// TIA Portal project "TNprojINZ" (V15.1)

(* hardware
DEVICE "S71500/ET200MP station_1"  S7-1500 station
   slot 0: "Rail_0"  Rack  6ES7 590-1***0-0AA0
   slot 1: "PLC_1"  CPU 1516-3 PN/DP  6ES7 516-3AN01-0AB0  V2.5
      slot 3: "CPU display_1"  6ES7591-1BA00-0AA0
   slot 2: "DI 32x24VDC HF_1"  DI 32x24VDC HF  6ES7 521-1BL00-0AB0  V2.1
   slot 3: "DQ 32x24VDC/0.5A ST_1"  DQ 32x24VDC/0.5A ST  6ES7 522-1BL00-0AB0  V2.0
   slot 4: "AI 8xU/I/RTD/TC ST_1"  AI 8xU/I/RTD/TC ST  6ES7 531-7KF00-0AB0  V2.0
   slot 5: "AQ 4xU/I ST_1"  AQ 4xU/I ST  6ES7 532-5HD00-0AB0  V2.0
DEVICE "HMI_1"  TP700 Comfort
   slot 0: "HMI_1"  TP700 Comfort  6AV2 124-0GC01-0AX0  15.1.0.0
   slot 1: "HMI_RT_1"  TP700 Comfort  6AV2 124-0GC01-0AX0  15.1.0.0
   slot 5: "HMI_1.IE_CP_1"  PROFINET Interface  15.0.1.0
      slot 1: "PROFINET Interface_1"  PROFINET Interface
         slot 1: "Port_1"  Port
         slot 2: "Port_2"  Port
   slot 7: "HMI_1.MPI/DP_CP_1"  MPI/DP Interface  15.0.1.0
*)

// ===== PLC "PLC_1"  CPU 1516-3 PN/DP =====

VAR_GLOBAL   // PLC tag table "Default tag table"
   "System_Byte" AT %MB1 : Byte;
   "FirstScan" AT %M1.0 : Bool;
   "DiagStatusUpdate" AT %M1.1 : Bool;
   "AlwaysTRUE" AT %M1.2 : Bool;
   "AlwaysFALSE" AT %M1.3 : Bool;
   "Clock_Byte" AT %MB0 : Byte;
   "Clock_10Hz" AT %M0.0 : Bool;
   "Clock_5Hz" AT %M0.1 : Bool;
   "Clock_2.5Hz" AT %M0.2 : Bool;
   "Clock_2Hz" AT %M0.3 : Bool;
   "Clock_1.25Hz" AT %M0.4 : Bool;
   "Clock_1Hz" AT %M0.5 : Bool;
   "Clock_0.625Hz" AT %M0.6 : Bool;
   "Clock_0.5Hz" AT %M0.7 : Bool;
   "Tag_1" AT %C3 : Counter;
END_VAR

DATA_BLOCK "Ster pompami"   // DB1
{ S7_Optimized_Access := 'TRUE' }
VERSION : 0.1
   VAR
      "przegrzana P1" : Bool;
      "przegrzana P2" : Bool;
      "przegrzana P3" : Bool;
      "przegrzana P4" : Bool;
      "przegrzana P5" : Bool;
      "przegrzana P6" : Bool;
      "przegrzana P7" : Bool;
      "przegrzana P8" : Bool;
   END_VAR
BEGIN
END_DATA_BLOCK

DATA_BLOCK "HMI komunikacja"   // DB2
{ S7_Optimized_Access := 'TRUE' }
VERSION : 0.1
   VAR
      "HMI Temp max Z1" : Real;   // zadany w HMI, następna part produktu
      "HMI Temp max Z2" : Real;   // zadany w HMI, następna part produktu
      "HMI Temp max Z3" : Real;   // zadany w HMI, następna part produktu
      "HMI Temp max Z4" : Real;   // zadany w HMI, następna part produktu
      "HMI poziom cieczy Z1" : Real;   // zadany w HMI, następna part produktu
      "HMI poziom cieczy Z2" : Real;   // zadany w HMI, następna part produktu
      "HMI poziom cieczy Z3" : Real;   // zadany w HMI, następna part produktu
      "HMI poziom cieczy Z4" : Real;   // zadany w HMI, następna part produktu
      "Czas utrz T w Z1 (timer)" : Real := 0.0;
      "Czas utrz T w Z2 (timer)" : Real := 0.0;
      "Czas utrz T w Z3 (timer)" : Real := 0.0;
      "Czas utrz T w Z4 (timer)" : Real := 0.0;
      "HMI czas utrz T  Z1" : Real := 0.0;   // zadany w HMI, następna part produktu
      "HMI czas utrz T  Z2" : Real := 0.0;   // zadany w HMI, następna part produktu
      "HMI czas utrz T  Z3" : Real := 0.0;   // zadany w HMI, następna part produktu
      "HMI czas utrz T  Z4" : Real := 0.0;   // zadany w HMI, następna part produktu
      "rura blue P5 i P6" : Bool := 0;
      "rura blue P1 i P2" : Bool := 0;
      "Start/Stop" : Bool := 0;
      "Blokada zmiany par. PRO" : Bool := 0;
   END_VAR
BEGIN
END_DATA_BLOCK

DATA_BLOCK "OPC - z LabVIEW"   // DB3
{ S7_Optimized_Access := 'FALSE' }
VERSION : 0.1
   VAR
      "Temp P1" : Real;
      "Temp P2" : Real;
      "Temp P3" : Real;
      "Temp P4" : Real;
      "Temp P5" : Real;
      "Temp P6" : Real;
      "Temp P7" : Real;
      "Temp P8" : Real;
      "Temp cieczy w zb1" : Real;
      "Temp cieczy w zb2" : Real;
      "Temp cieczy w zb3" : Real;
      "Temp cieczy w zb4" : Real;
      "Poziom zbiornik 1" : Real;
      "Poziom zbiornik 2" : Real;
      "Poziom zbiornik 3" : Real;
      "Poziom zbiornik 4" : Real;
      komTESTz : Bool := 0;
   END_VAR
BEGIN
END_DATA_BLOCK

DATA_BLOCK "OPC - do LabVIEW"   // DB4
{ S7_Optimized_Access := 'FALSE' }
VERSION : 0.1
   VAR
      "PRO Temp max Z1" : Real;   // dla SFC, aktualna partia produktu
      "PRO Temp max Z2" : Real;   // dla SFC, aktualna partia produktu
      "PRO Temp max Z3" : Real;   // dla SFC, aktualna partia produktu
      "PRO Temp max Z4" : Real;   // dla SFC, aktualna partia produktu
      "PRO poziom cieczy Z1" : Real;   // dla SFC, aktualna partia produktu
      "PRO poziom cieczy Z2" : Real;   // dla SFC, aktualna partia produktu
      "PRO poziom cieczy Z3" : Real;   // dla SFC, aktualna partia produktu
      "PRO poziom cieczy Z4" : Real;   // dla SFC, aktualna partia produktu
      "PRO czas utrz T  Z1" : Real := 0.0;   // dla SFC, aktualna partia produktu
      "PRO czas utrz T  Z2" : Real := 0.0;   // dla SFC, aktualna partia produktu
      "PRO czas utrz T  Z3" : Real := 0.0;   // dla SFC, aktualna partia produktu
      "PRO czas utrz T  Z4" : Real := 0.0;   // dla SFC, aktualna partia produktu
      Awaria : Bool := 0;
      "Pompa 1" : Bool := 0;
      "Pompa 2" : Bool := 0;
      "Pompa 3" : Bool := 0;
      "Pompa 4" : Bool := 0;
      "Pompa 5" : Bool := 0;
      "Pompa 6" : Bool := 0;
      "Pompa 7" : Bool := 0;
      "Pompa 8" : Bool := 0;
      "Zawór wlotowy 1" : Bool := 0;
      "Zawór wlotowy 2" : Bool := 0;
      "Zawór wlotowy 3" : Bool := 0;
      "Grzałka 1" : Bool := 0;
      "Grzałka 2" : Bool := 0;
      "Grzałka 3" : Bool := 0;
      "Grzałka 4" : Bool := 0;
      "HMI konserwacja P1" : Bool := 0;
      "HMI konserwacja P2" : Bool := 0;
      "HMI konserwacja P3" : Bool := 0;
      "HMI konserwacja P4" : Bool := 0;
      "HMI konserwacja P5" : Bool := 0;
      "HMI konserwacja P6" : Bool := 0;
      "HMI konserwacja P7" : Bool := 0;
      "HMI konserwacja P8" : Bool := 0;
      "Zawór spustowy Z1" : Bool := 0;
      "Zawór spustowy Z2" : Bool := 0;
      "Zawór spustowy Z3" : Bool := 0;
      "Zawór spustowy Z4" : Bool := 0;
      komTESTdo : Bool := 0;
   END_VAR
BEGIN
END_DATA_BLOCK

DATA_BLOCK "Ster grzałki/zbior"   // DB5
{ S7_Optimized_Access := 'TRUE' }
VERSION : 0.1
   VAR
      HISTgrzałka1 : Bool;
      HISTgrzałka2 : Bool;
      HISTgrzałka3 : Bool;
      HISTgrzałka4 : Bool;
      "Wszystkie zbiorniki puste" : Bool;
      "Z1 opróżniony" : Bool;
      "Z2 opróżniony" : Bool;
      "Z3 opróżniony" : Bool;
   END_VAR
BEGIN
END_DATA_BLOCK

// folder: DB - Instance

DATA_BLOCK "Zbiornik 1_DB"   // DB6
{ S7_Optimized_Access := 'TRUE' }
VERSION : 0.1
// stored: InstanceOfName Zbiornik 1
"Zbiornik 1"
BEGIN
END_DATA_BLOCK

DATA_BLOCK "Zbiornik 2_DB"   // DB15
{ S7_Optimized_Access := 'TRUE' }
VERSION : 0.1
// stored: InstanceOfName Zbiornik 2
"Zbiornik 2"
BEGIN
END_DATA_BLOCK

DATA_BLOCK "Zbiornik 3_DB"   // DB16
{ S7_Optimized_Access := 'TRUE' }
VERSION : 0.1
// stored: InstanceOfName Zbiornik 3
"Zbiornik 3"
BEGIN
END_DATA_BLOCK

DATA_BLOCK "Zbiornik 4_DB"   // DB17
{ S7_Optimized_Access := 'TRUE' }
VERSION : 0.1
// stored: InstanceOfName Zbiornik 4
"Zbiornik 4"
BEGIN
END_DATA_BLOCK

DATA_BLOCK "SCL - Sterowanie pompami_DB"   // DB18
{ S7_Optimized_Access := 'TRUE' }
VERSION : 0.1
// stored: InstanceOfName SCL - Sterowanie pompami
"SCL - Sterowanie pompami"
BEGIN
END_DATA_BLOCK

DATA_BLOCK "SCL - Napełnianie i kontrola_DB"   // DB19
{ S7_Optimized_Access := 'TRUE' }
VERSION : 0.1
// stored: InstanceOfName SCL - Napełnianie i kontrola
"SCL - Napełnianie i kontrola"
BEGIN
END_DATA_BLOCK

DATA_BLOCK "SCL - Grzanie_DB"   // DB20
{ S7_Optimized_Access := 'TRUE' }
VERSION : 0.1
// stored: InstanceOfName SCL - Grzanie
"SCL - Grzanie"
BEGIN
END_DATA_BLOCK

DATA_BLOCK "SCL - Awaria_DB"   // DB21
{ S7_Optimized_Access := 'TRUE' }
VERSION : 0.1
// stored: InstanceOfName SCL - Awaria i zabezpieczenia par.
"SCL - Awaria i zabezpieczenia par."
BEGIN
END_DATA_BLOCK

DATA_BLOCK "FB - pompy_DB"   // DB22
{ S7_Optimized_Access := 'TRUE' }
VERSION : 0.1
// stored: InstanceOfName FB - pompy
"FB - pompy"
BEGIN
END_DATA_BLOCK

DATA_BLOCK "FB - grzałki_DB"   // DB23
{ S7_Optimized_Access := 'TRUE' }
VERSION : 0.1
// stored: InstanceOfName FB - grzałki
"FB - grzałki"
BEGIN
END_DATA_BLOCK

// folder: System blocks/Program resources

DATA_BLOCK "IEC_Timer_2_DB"   // DB7
{ S7_Optimized_Access := 'TRUE' }
AUTHOR : Simatic
FAMILY : IEC
NAME : IEC_TMR
VERSION : 1.0
// stored: InstanceOfName IEC_TIMER
"IEC_TIMER"
BEGIN
END_DATA_BLOCK

DATA_BLOCK "IEC_Timer_3_DB"   // DB12
{ S7_Optimized_Access := 'TRUE' }
AUTHOR : Simatic
FAMILY : IEC
NAME : IEC_TMR
VERSION : 1.0
// stored: InstanceOfName IEC_TIMER
"IEC_TIMER"
BEGIN
END_DATA_BLOCK

DATA_BLOCK "IEC_Timer_1_DB"   // DB13
{ S7_Optimized_Access := 'TRUE' }
AUTHOR : Simatic
FAMILY : IEC
NAME : IEC_TMR
VERSION : 1.0
// stored: InstanceOfName IEC_TIMER
"IEC_TIMER"
BEGIN
END_DATA_BLOCK

DATA_BLOCK "IEC_Timer_4_DB"   // DB14
{ S7_Optimized_Access := 'TRUE' }
AUTHOR : Simatic
FAMILY : IEC
NAME : IEC_TMR
VERSION : 1.0
// stored: InstanceOfName IEC_TIMER
"IEC_TIMER"
BEGIN
END_DATA_BLOCK

DATA_BLOCK "IEC_Timer_0_DB"   // DB24
{ S7_Optimized_Access := 'TRUE' }
AUTHOR : Simatic
FAMILY : IEC
NAME : IEC_TMR
VERSION : 1.0
// stored: InstanceOfName IEC_TIMER
"IEC_TIMER"
BEGIN
END_DATA_BLOCK

DATA_BLOCK "IEC_Timer_0_DB_2"   // DB26
{ S7_Optimized_Access := 'TRUE' }
AUTHOR : Simatic
FAMILY : IEC
NAME : IEC_TMR
VERSION : 1.0
// stored: InstanceOfName IEC_TIMER
"IEC_TIMER"
BEGIN
END_DATA_BLOCK

// folder: Zbiorniki - globalne

DATA_BLOCK "Z1 globalne"   // DB8
{ S7_Optimized_Access := 'TRUE' }
VERSION : 0.1
   VAR
      "Czy Z1 pełny?" : Bool := 0;
      "Ciecz Z1 nagrzana" : Bool;
      "awaria Z1 sfc" : Bool;
      "grzanie Z1 sfc" : Bool;
      "napełnianie Z1 sfc" : Bool;
      "opróżnianie Z1 sfc" : Bool;
      "Z1 gotowy" : Bool;
      "Awaria reset sfc Z1" : Bool;
      "Z1 opóźnienie" : Bool;
   END_VAR
BEGIN
END_DATA_BLOCK

DATA_BLOCK "Z2 globalne"   // DB9
{ S7_Optimized_Access := 'TRUE' }
VERSION : 0.1
   VAR
      "Czy Z2 pełny?" : Bool;
      "Ciecz Z2 nagrzana" : Bool;
      "awaria Z2 sfc" : Bool;
      "grzanie Z2 sfc" : Bool;
      "napełnianie Z2 sfc" : Bool;
      "opróżnianie Z2 sfc" : Bool;
      "Z2 gotowy" : Bool;
      "Awaria reset sfc Z2" : Bool;
      "Z2 opóźnienie" : Bool;
   END_VAR
BEGIN
END_DATA_BLOCK

DATA_BLOCK "Z3 globalne"   // DB10
{ S7_Optimized_Access := 'TRUE' }
VERSION : 0.1
   VAR
      "Czy Z3 pełny?" : Bool;
      "Ciecz Z3 nagrzana" : Bool;
      "awaria Z3 sfc" : Bool;
      "grzanie Z3 sfc" : Bool;
      "napełnianie Z3 sfc" : Bool;
      "opróżnianie Z3 sfc" : Bool;
      "Z3 gotowy" : Bool;
      "Awaria reset sfc Z3" : Bool;
      "Z3 opóźnienie" : Bool;
   END_VAR
BEGIN
END_DATA_BLOCK

DATA_BLOCK "Z4 globalne"   // DB11
{ S7_Optimized_Access := 'TRUE' }
VERSION : 0.1
   VAR
      "Czy Z4 pełny?" : Bool;
      "Ciecz Z4 nagrzana" : Bool;
      "awaria Z4 sfc" : Bool;
      "grzanie Z4 sfc" : Bool;
      "napełnianie Z4 sfc" : Bool;
      "opróżnianie Z4 sfc" : Bool;
      "Z4 gotowy" : Bool;
      "Awaria reset sfc Z4" : Bool;
   END_VAR
BEGIN
END_DATA_BLOCK

// folder: (top level)

FUNCTION_BLOCK "Zbiornik 1"   // FB1, GRAPH_PLUS
{ S7_Optimized_Access := 'TRUE' }
VERSION : 0.1
   VAR_INPUT
      OFF_SQ : Bool := false;   // Turn sequence off
      INIT_SQ : Bool := false;   // Set sequence to initial state
      ACK_EF : Bool := false;   // Acknowledge all errors and faults
      S_PREV : Bool := false;   // Output previous step in parameter S_NO
      S_NEXT : Bool := false;   // Indicate next step in parameter S_NO
      SW_AUTO : Bool := false;   // Automatic mode
      SW_TAP : Bool := false;   // Semiautomatic/switch with transition
      SW_TOP : Bool := false;   // Semiautomatic/ignore transition
      SW_MAN : Bool := false;   // Manual mode
      S_SEL : Int := 0;   // Select step to be output to S_NO
      S_ON : Bool := false;   // Activate step indicated in S_NO
      S_OFF : Bool := false;   // Deactivate step indicated S_NO
      T_PUSH : Bool := false;   // Enable transition to switch in semi automatic mode
   END_VAR
   VAR_OUTPUT
      S_NO : Int := 0;   // Step number
      S_MORE : Bool := false;   // More steps are available and can be shown in S_NO
      S_ACTIVE : Bool := false;   // Step indicated in S_NO is active
      ERR_FLT : Bool := false;   // Interlock or supervision group error
      AUTO_ON : Bool := false;   // Automatic mode is active
      TAP_ON : Bool := false;   // Semiautomatic mode/step with transition enabled
      TOP_ON : Bool := false;   // Semiautomatic mode/ignore transition enabled
      MAN_ON : Bool := false;   // Manual mode is active
   END_VAR
   VAR
      HMI_INFO : Array[0..10] of UInt;
      IF_PAR : G7_IfParPlus_V6;
      RT_DATA : G7_RTDataPlus_V6;   // Internal data area
      "Start/stop" : G7_TransitionPlus_V6;   // Transition structure
      "Start/stop1" : G7_TransitionPlus_V6;   // Transition structure
      "Czy pełny?" : G7_TransitionPlus_V6;   // Transition structure
      "Gotowy?" : G7_TransitionPlus_V6;   // Transition structure
      "Czy pusty?" : G7_TransitionPlus_V6;   // Transition structure
      Wznowienie : G7_TransitionPlus_V6;   // Transition structure
      Trans9 : G7_TransitionPlus_V6;   // Transition structure
      Trans10 : G7_TransitionPlus_V6;   // Transition structure
      Init : G7_StepPlus_V6;   // Step structure
      "reset/kontrola" : G7_StepPlus_V6;   // Step structure
      Napełnianie : G7_StepPlus_V6;   // Step structure
      Grzanie : G7_StepPlus_V6;   // Step structure
      Opróżnianie : G7_StepPlus_V6;   // Step structure
      "Awaria HMI" : G7_StepPlus_V6;   // Step structure
      Opóźnienie : G7_StepPlus_V6;   // Step structure
      Step12 : G7_StepPlus_V6;   // Step structure
      SINI : Array[0..3] of USInt;
      LSTT : Array[0..7] of USInt;
      ATAJ : Array[0..7] of USInt;
      ATAB : Array[0..7] of USInt;
      PSTT : Array[0..7] of USInt;
      NSTT : Array[0..7] of USInt;
      ASSJ : Array[0..7] of USInt;
      ASSB : Array[0..7] of USInt;
      PTTS : Array[0..7] of USInt;
      NTTS : Array[0..7] of USInt;
      SW_SQTS : Array[0..7] of USInt;
      SWITCH : Array[0..1] of USInt;
      TVX : Array[0..3] of USInt;
      TTX : Array[0..3] of USInt;
      TSX : Array[0..3] of USInt;
      S00X : Array[0..3] of USInt;
      SOFFX : Array[0..3] of USInt;
      SONX : Array[0..3] of USInt;
      SAX : Array[0..3] of USInt;
      SERRX : Array[0..8] of USInt;
      SMX : Array[0..8] of USInt;
      S0X : Array[0..8] of USInt;
      S1X : Array[0..8] of USInt;
      IL_ALARM_INST : Diag_Alarm;
      SUP_ALARM_INST : Diag_Alarm;
      STEP_TIME_ALARM_INST : Diag_Alarm;
      IEC_TIMER_INST : IEC_TIMER;
      TRANSACTION_FLAG : Bool := false;
   END_VAR
   // SINI[0] := 2;
   // SINI[2] := 255;
   // SINI[3] := 255;
   // LSTT[0] := 255;
   // LSTT[1] := 255;
   // LSTT[2] := 255;
   // LSTT[3] := 255;
   // LSTT[4] := 255;
   // LSTT[5] := 1;
   // ATAJ[1] := 1;
   // ATAJ[2] := 2;
   // ATAJ[3] := 3;
   // ATAJ[4] := 4;
   // ATAJ[5] := 5;
   // ATAB[1] := 1;
   // ATAB[2] := 2;
   // ATAB[3] := 3;
   // ATAB[4] := 4;
   // ATAB[5] := 5;
   // PSTT[1] := 1;
   // PSTT[2] := 2;
   // PSTT[3] := 3;
   // PSTT[4] := 4;
   // PSTT[5] := 5;
   // NSTT[0] := 1;
   // NSTT[1] := 2;
   // NSTT[2] := 3;
   // NSTT[3] := 4;
   // NSTT[4] := 6;
   // NSTT[5] := 1;
   // ASSJ[1] := 1;
   // ASSJ[2] := 2;
   // ASSJ[3] := 3;
   // ASSJ[4] := 4;
   // ASSJ[5] := 5;
   // ASSB[1] := 1;
   // ASSB[2] := 5;
   // ASSB[3] := 3;
   // ASSB[4] := 4;
   // ASSB[5] := 2;
   // PTTS[0] := 255;
   // PTTS[2] := 1;
   // PTTS[3] := 2;
   // PTTS[4] := 3;
   // PTTS[5] := 1;
   // NTTS[1] := 1;
   // NTTS[2] := 2;
   // NTTS[3] := 3;
   // NTTS[4] := 4;
   // NTTS[5] := 5;
   // SW_SQTS[2] := 1;
   // SW_SQTS[3] := 1;
   // SW_SQTS[4] := 1;
   // SW_SQTS[5] := 2;
   // SWITCH[0] := 160;
   // TVX[0] := 16#1;
   // TTX[0] := 16#1;
   // TSX[0] := 16#1;
   // S00X[0] := 16#1;
   // SOFFX[0] := 16#1;
   // SONX[0] := 16#1;
   // SAX[0] := 16#1;
   // SERRX[0] := 16#1;
   // SMX[0] := 16#1;
   // S0X[0] := 16#1;
   // S1X[0] := 16#1;
   // LSTT[6] := 255;
   // ATAJ[6] := 6;
   // ATAB[6] := 6;
   // PSTT[6] := 6;
   // NSTT[6] := 7;
   // ASSJ[6] := 6;
   // ASSB[6] := 6;
   // PTTS[6] := 4;
   // NTTS[6] := 6;
   // SW_SQTS[6] := 1;
   // LSTT[7] := 1;
   // ATAJ[7] := 7;
   // ATAB[7] := 7;
   // PSTT[7] := 7;
   // NSTT[7] := 1;
   // ASSJ[7] := 7;
   // ASSB[7] := 7;
   // PTTS[7] := 6;
   // NTTS[7] := 7;
   // SW_SQTS[7] := 1;
BEGIN
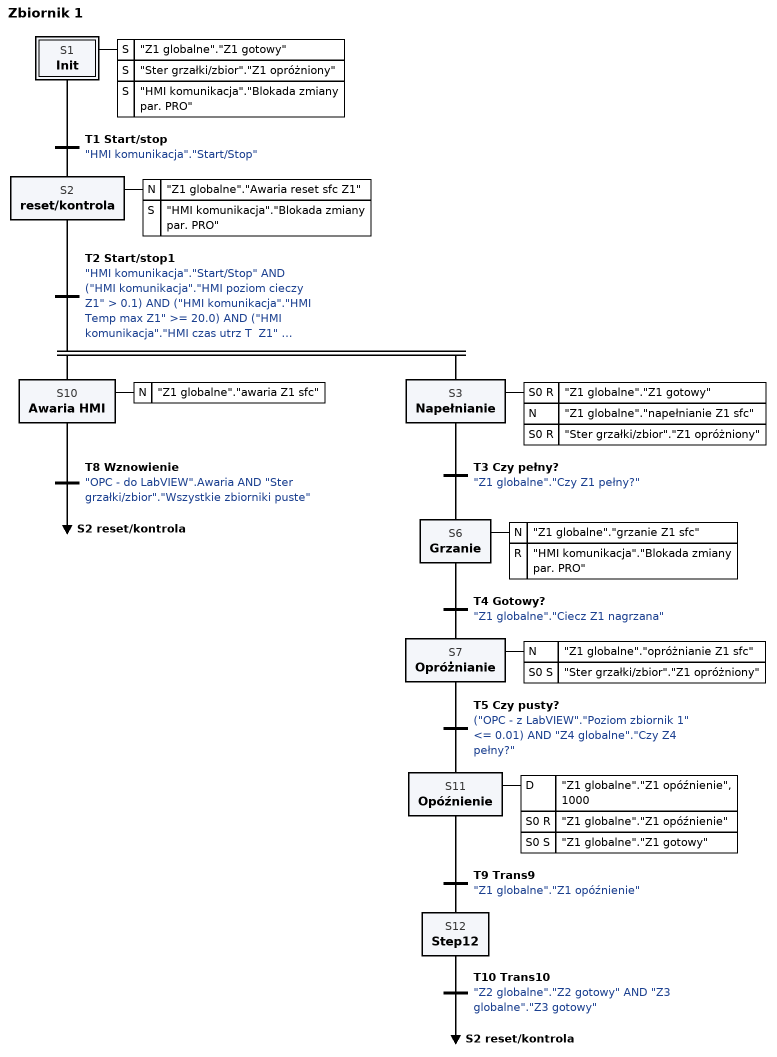
   // sequencer 1
   INITIAL_STEP Init:   // S1, max time T#10S, warning time T#7S
              S    "Z1 globalne"."Z1 gotowy"
              S    "Ster grzałki/zbior"."Z1 opróżniony"
              S    "HMI komunikacja"."Blokada zmiany par. PRO"
   END_STEP
   TRANSITION "Start/stop" FROM Init TO "reset/kontrola"   // T1
      := "HMI komunikacja"."Start/Stop";
   END_TRANSITION
   STEP "reset/kontrola":   // S2, max time T#10S, warning time T#7S
              N    "Z1 globalne"."Awaria reset sfc Z1"
              S    "HMI komunikacja"."Blokada zmiany par. PRO"
   END_STEP
   TRANSITION "Start/stop1" FROM "reset/kontrola" TO ("Awaria HMI", Napełnianie)   // T2
      := "HMI komunikacja"."Start/Stop" AND ("HMI komunikacja"."HMI poziom cieczy Z1" > 0.1) AND ("HMI komunikacja"."HMI Temp max Z1" >= 20.0) AND ("HMI komunikacja"."HMI czas utrz T  Z1" > 0.1) AND "Z2 globalne"."Z2 gotowy" AND "Z3 globalne"."Z3 gotowy";
   END_TRANSITION
   STEP Napełnianie:   // S3, max time T#10S, warning time T#7S
          S0  R    "Z1 globalne"."Z1 gotowy"
              N    "Z1 globalne"."napełnianie Z1 sfc"
          S0  R    "Ster grzałki/zbior"."Z1 opróżniony"
   END_STEP
   TRANSITION "Czy pełny?" FROM Napełnianie TO Grzanie   // T3
      := "Z1 globalne"."Czy Z1 pełny?";
   END_TRANSITION
   STEP Grzanie:   // S6, max time T#10S, warning time T#7S
              N    "Z1 globalne"."grzanie Z1 sfc"
              R    "HMI komunikacja"."Blokada zmiany par. PRO"
   END_STEP
   TRANSITION "Gotowy?" FROM Grzanie TO Opróżnianie   // T4
      := "Z1 globalne"."Ciecz Z1 nagrzana";
   END_TRANSITION
   STEP Opróżnianie:   // S7, max time T#10S, warning time T#7S
              N    "Z1 globalne"."opróżnianie Z1 sfc"
          S0  S    "Ster grzałki/zbior"."Z1 opróżniony"
   END_STEP
   TRANSITION "Czy pusty?" FROM Opróżnianie TO Opóźnienie   // T5
      := ("OPC - z LabVIEW"."Poziom zbiornik 1" <= 0.01) AND "Z4 globalne"."Czy Z4 pełny?";
   END_TRANSITION
   STEP "Awaria HMI":   // S10, max time T#10S, warning time T#7S
              N    "Z1 globalne"."awaria Z1 sfc"
   END_STEP
   TRANSITION Wznowienie FROM "Awaria HMI" TO "reset/kontrola"   // T8, jump
      := "OPC - do LabVIEW".Awaria AND "Ster grzałki/zbior"."Wszystkie zbiorniki puste";
   END_TRANSITION
   STEP Opóźnienie:   // S11, max time T#10S, warning time T#7S
              D    "Z1 globalne"."Z1 opóźnienie", 1000
          S0  R    "Z1 globalne"."Z1 opóźnienie"
          S0  S    "Z1 globalne"."Z1 gotowy"
   END_STEP
   TRANSITION Trans9 FROM Opóźnienie TO Step12   // T9
      := "Z1 globalne"."Z1 opóźnienie";
   END_TRANSITION
   STEP Step12:   // S12, max time T#10S, warning time T#7S
   END_STEP
   TRANSITION Trans10 FROM Step12 TO "reset/kontrola"   // T10, jump
      := "Z2 globalne"."Z2 gotowy" AND "Z3 globalne"."Z3 gotowy";
   END_TRANSITION
END_FUNCTION_BLOCK

FUNCTION_BLOCK "Zbiornik 2"   // FB2, GRAPH_PLUS
{ S7_Optimized_Access := 'TRUE' }
VERSION : 0.1
   VAR_INPUT
      OFF_SQ : Bool := false;   // Turn sequence off
      INIT_SQ : Bool := false;   // Set sequence to initial state
      ACK_EF : Bool := false;   // Acknowledge all errors and faults
      S_PREV : Bool := false;   // Output previous step in parameter S_NO
      S_NEXT : Bool := false;   // Indicate next step in parameter S_NO
      SW_AUTO : Bool := false;   // Automatic mode
      SW_TAP : Bool := false;   // Semiautomatic/switch with transition
      SW_TOP : Bool := false;   // Semiautomatic/ignore transition
      SW_MAN : Bool := false;   // Manual mode
      S_SEL : Int := 0;   // Select step to be output to S_NO
      S_ON : Bool := false;   // Activate step indicated in S_NO
      S_OFF : Bool := false;   // Deactivate step indicated S_NO
      T_PUSH : Bool := false;   // Enable transition to switch in semi automatic mode
   END_VAR
   VAR_OUTPUT
      S_NO : Int := 0;   // Step number
      S_MORE : Bool := false;   // More steps are available and can be shown in S_NO
      S_ACTIVE : Bool := false;   // Step indicated in S_NO is active
      ERR_FLT : Bool := false;   // Interlock or supervision group error
      AUTO_ON : Bool := false;   // Automatic mode is active
      TAP_ON : Bool := false;   // Semiautomatic mode/step with transition enabled
      TOP_ON : Bool := false;   // Semiautomatic mode/ignore transition enabled
      MAN_ON : Bool := false;   // Manual mode is active
   END_VAR
   VAR
      HMI_INFO : Array[0..10] of UInt;
      IF_PAR : G7_IfParPlus_V6;
      RT_DATA : G7_RTDataPlus_V6;   // Internal data area
      "Start/stop" : G7_TransitionPlus_V6;   // Transition structure
      "Start/stop1" : G7_TransitionPlus_V6;   // Transition structure
      "Czy_pełny?" : G7_TransitionPlus_V6;   // Transition structure
      "Gotowy?" : G7_TransitionPlus_V6;   // Transition structure
      "Czy_pusty?" : G7_TransitionPlus_V6;   // Transition structure
      Wznowienie : G7_TransitionPlus_V6;   // Transition structure
      Trans9 : G7_TransitionPlus_V6;   // Transition structure
      Trans10 : G7_TransitionPlus_V6;   // Transition structure
      Init : G7_StepPlus_V6;   // Step structure
      "reset/kontrola" : G7_StepPlus_V6;   // Step structure
      Napełnianie : G7_StepPlus_V6;   // Step structure
      Grzanie : G7_StepPlus_V6;   // Step structure
      Opróżnianie : G7_StepPlus_V6;   // Step structure
      "Awaria HMI" : G7_StepPlus_V6;   // Step structure
      Opóźnienie : G7_StepPlus_V6;   // Step structure
      Step12 : G7_StepPlus_V6;   // Step structure
      SINI : Array[0..3] of USInt;
      LSTT : Array[0..7] of USInt;
      ATAJ : Array[0..7] of USInt;
      ATAB : Array[0..7] of USInt;
      PSTT : Array[0..7] of USInt;
      NSTT : Array[0..7] of USInt;
      ASSJ : Array[0..7] of USInt;
      ASSB : Array[0..7] of USInt;
      PTTS : Array[0..7] of USInt;
      NTTS : Array[0..7] of USInt;
      SW_SQTS : Array[0..7] of USInt;
      SWITCH : Array[0..1] of USInt;
      TVX : Array[0..3] of USInt;
      TTX : Array[0..3] of USInt;
      TSX : Array[0..3] of USInt;
      S00X : Array[0..3] of USInt;
      SOFFX : Array[0..3] of USInt;
      SONX : Array[0..3] of USInt;
      SAX : Array[0..3] of USInt;
      SERRX : Array[0..8] of USInt;
      SMX : Array[0..8] of USInt;
      S0X : Array[0..8] of USInt;
      S1X : Array[0..8] of USInt;
      IL_ALARM_INST : Diag_Alarm;
      SUP_ALARM_INST : Diag_Alarm;
      STEP_TIME_ALARM_INST : Diag_Alarm;
      IEC_TIMER_INST : IEC_TIMER;
      TRANSACTION_FLAG : Bool := false;
   END_VAR
   // SINI[0] := 2;
   // SINI[2] := 255;
   // SINI[3] := 255;
   // LSTT[0] := 255;
   // LSTT[1] := 255;
   // LSTT[2] := 255;
   // LSTT[3] := 255;
   // LSTT[4] := 255;
   // LSTT[5] := 1;
   // ATAJ[1] := 1;
   // ATAJ[2] := 2;
   // ATAJ[3] := 3;
   // ATAJ[4] := 4;
   // ATAJ[5] := 5;
   // ATAB[1] := 1;
   // ATAB[2] := 2;
   // ATAB[3] := 3;
   // ATAB[4] := 4;
   // ATAB[5] := 5;
   // PSTT[1] := 1;
   // PSTT[2] := 2;
   // PSTT[3] := 3;
   // PSTT[4] := 4;
   // PSTT[5] := 5;
   // NSTT[0] := 1;
   // NSTT[1] := 2;
   // NSTT[2] := 3;
   // NSTT[3] := 4;
   // NSTT[4] := 6;
   // NSTT[5] := 1;
   // ASSJ[1] := 1;
   // ASSJ[2] := 2;
   // ASSJ[3] := 3;
   // ASSJ[4] := 4;
   // ASSJ[5] := 5;
   // ASSB[1] := 1;
   // ASSB[2] := 5;
   // ASSB[3] := 3;
   // ASSB[4] := 4;
   // ASSB[5] := 2;
   // PTTS[0] := 255;
   // PTTS[2] := 1;
   // PTTS[3] := 2;
   // PTTS[4] := 3;
   // PTTS[5] := 1;
   // NTTS[1] := 1;
   // NTTS[2] := 2;
   // NTTS[3] := 3;
   // NTTS[4] := 4;
   // NTTS[5] := 5;
   // SW_SQTS[2] := 1;
   // SW_SQTS[3] := 1;
   // SW_SQTS[4] := 1;
   // SW_SQTS[5] := 2;
   // SWITCH[0] := 160;
   // TVX[0] := 16#1;
   // TTX[0] := 16#1;
   // TSX[0] := 16#1;
   // S00X[0] := 16#1;
   // SOFFX[0] := 16#1;
   // SONX[0] := 16#1;
   // SAX[0] := 16#1;
   // SERRX[0] := 16#1;
   // SMX[0] := 16#1;
   // S0X[0] := 16#1;
   // S1X[0] := 16#1;
   // LSTT[6] := 255;
   // ATAJ[6] := 6;
   // ATAB[6] := 6;
   // PSTT[6] := 6;
   // NSTT[6] := 7;
   // ASSJ[6] := 6;
   // ASSB[6] := 6;
   // PTTS[6] := 4;
   // NTTS[6] := 6;
   // SW_SQTS[6] := 1;
   // LSTT[7] := 1;
   // ATAJ[7] := 7;
   // ATAB[7] := 7;
   // PSTT[7] := 7;
   // NSTT[7] := 1;
   // ASSJ[7] := 7;
   // ASSB[7] := 7;
   // PTTS[7] := 6;
   // NTTS[7] := 7;
   // SW_SQTS[7] := 1;
BEGIN
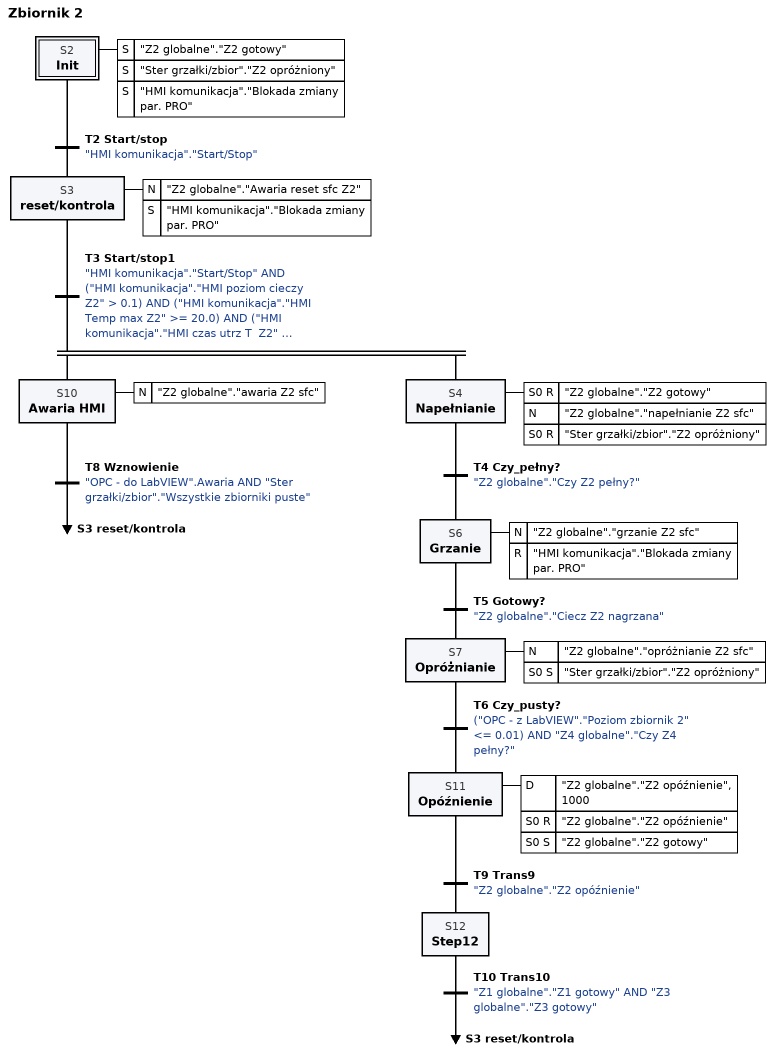
   // sequencer 1
   INITIAL_STEP Init:   // S2, max time T#10S, warning time T#7S
              S    "Z2 globalne"."Z2 gotowy"
              S    "Ster grzałki/zbior"."Z2 opróżniony"
              S    "HMI komunikacja"."Blokada zmiany par. PRO"
   END_STEP
   TRANSITION "Start/stop" FROM Init TO "reset/kontrola"   // T2
      := "HMI komunikacja"."Start/Stop";
   END_TRANSITION
   STEP "reset/kontrola":   // S3, max time T#10S, warning time T#7S
              N    "Z2 globalne"."Awaria reset sfc Z2"
              S    "HMI komunikacja"."Blokada zmiany par. PRO"
   END_STEP
   TRANSITION "Start/stop1" FROM "reset/kontrola" TO ("Awaria HMI", Napełnianie)   // T3
      := "HMI komunikacja"."Start/Stop" AND ("HMI komunikacja"."HMI poziom cieczy Z2" > 0.1) AND ("HMI komunikacja"."HMI Temp max Z2" >= 20.0) AND ("HMI komunikacja"."HMI czas utrz T  Z2" > 0.1) AND "Z1 globalne"."Z1 gotowy" AND "Z3 globalne"."Z3 gotowy";
   END_TRANSITION
   STEP Napełnianie:   // S4, max time T#10S, warning time T#7S
          S0  R    "Z2 globalne"."Z2 gotowy"
              N    "Z2 globalne"."napełnianie Z2 sfc"
          S0  R    "Ster grzałki/zbior"."Z2 opróżniony"
   END_STEP
   TRANSITION "Czy_pełny?" FROM Napełnianie TO Grzanie   // T4
      := "Z2 globalne"."Czy Z2 pełny?";
   END_TRANSITION
   STEP Grzanie:   // S6, max time T#10S, warning time T#7S
              N    "Z2 globalne"."grzanie Z2 sfc"
              R    "HMI komunikacja"."Blokada zmiany par. PRO"
   END_STEP
   TRANSITION "Gotowy?" FROM Grzanie TO Opróżnianie   // T5
      := "Z2 globalne"."Ciecz Z2 nagrzana";
   END_TRANSITION
   STEP Opróżnianie:   // S7, max time T#10S, warning time T#7S
              N    "Z2 globalne"."opróżnianie Z2 sfc"
          S0  S    "Ster grzałki/zbior"."Z2 opróżniony"
   END_STEP
   TRANSITION "Czy_pusty?" FROM Opróżnianie TO Opóźnienie   // T6
      := ("OPC - z LabVIEW"."Poziom zbiornik 2" <= 0.01) AND "Z4 globalne"."Czy Z4 pełny?";
   END_TRANSITION
   STEP "Awaria HMI":   // S10, max time T#10S, warning time T#7S
              N    "Z2 globalne"."awaria Z2 sfc"
   END_STEP
   TRANSITION Wznowienie FROM "Awaria HMI" TO "reset/kontrola"   // T8, jump
      := "OPC - do LabVIEW".Awaria AND "Ster grzałki/zbior"."Wszystkie zbiorniki puste";
   END_TRANSITION
   STEP Opóźnienie:   // S11, max time T#10S, warning time T#7S
              D    "Z2 globalne"."Z2 opóźnienie", 1000
          S0  R    "Z2 globalne"."Z2 opóźnienie"
          S0  S    "Z2 globalne"."Z2 gotowy"
   END_STEP
   TRANSITION Trans9 FROM Opóźnienie TO Step12   // T9
      := "Z2 globalne"."Z2 opóźnienie";
   END_TRANSITION
   STEP Step12:   // S12, max time T#10S, warning time T#7S
   END_STEP
   TRANSITION Trans10 FROM Step12 TO "reset/kontrola"   // T10, jump
      := "Z1 globalne"."Z1 gotowy" AND "Z3 globalne"."Z3 gotowy";
   END_TRANSITION
END_FUNCTION_BLOCK

FUNCTION_BLOCK "Zbiornik 3"   // FB3, GRAPH_PLUS
{ S7_Optimized_Access := 'TRUE' }
VERSION : 0.1
   VAR_INPUT
      OFF_SQ : Bool := false;   // Turn sequence off
      INIT_SQ : Bool := false;   // Set sequence to initial state
      ACK_EF : Bool := false;   // Acknowledge all errors and faults
      S_PREV : Bool := false;   // Output previous step in parameter S_NO
      S_NEXT : Bool := false;   // Indicate next step in parameter S_NO
      SW_AUTO : Bool := false;   // Automatic mode
      SW_TAP : Bool := false;   // Semiautomatic/switch with transition
      SW_TOP : Bool := false;   // Semiautomatic/ignore transition
      SW_MAN : Bool := false;   // Manual mode
      S_SEL : Int := 0;   // Select step to be output to S_NO
      S_ON : Bool := false;   // Activate step indicated in S_NO
      S_OFF : Bool := false;   // Deactivate step indicated S_NO
      T_PUSH : Bool := false;   // Enable transition to switch in semi automatic mode
   END_VAR
   VAR_OUTPUT
      S_NO : Int := 0;   // Step number
      S_MORE : Bool := false;   // More steps are available and can be shown in S_NO
      S_ACTIVE : Bool := false;   // Step indicated in S_NO is active
      ERR_FLT : Bool := false;   // Interlock or supervision group error
      AUTO_ON : Bool := false;   // Automatic mode is active
      TAP_ON : Bool := false;   // Semiautomatic mode/step with transition enabled
      TOP_ON : Bool := false;   // Semiautomatic mode/ignore transition enabled
      MAN_ON : Bool := false;   // Manual mode is active
   END_VAR
   VAR
      HMI_INFO : Array[0..10] of UInt;
      IF_PAR : G7_IfParPlus_V6;
      RT_DATA : G7_RTDataPlus_V6;   // Internal data area
      "Start/stop" : G7_TransitionPlus_V6;   // Transition structure
      "Start/stop1" : G7_TransitionPlus_V6;   // Transition structure
      "Czy_pełny?" : G7_TransitionPlus_V6;   // Transition structure
      "Gotowy?" : G7_TransitionPlus_V6;   // Transition structure
      "Czy_pusty?" : G7_TransitionPlus_V6;   // Transition structure
      Wznowienie : G7_TransitionPlus_V6;   // Transition structure
      Trans9 : G7_TransitionPlus_V6;   // Transition structure
      Trans10 : G7_TransitionPlus_V6;   // Transition structure
      Init : G7_StepPlus_V6;   // Step structure
      "reset/kontrola" : G7_StepPlus_V6;   // Step structure
      Napełnianie : G7_StepPlus_V6;   // Step structure
      Grzanie : G7_StepPlus_V6;   // Step structure
      Opróżnianie : G7_StepPlus_V6;   // Step structure
      "Awaria HMI" : G7_StepPlus_V6;   // Step structure
      Opóźnienie : G7_StepPlus_V6;   // Step structure
      Step12 : G7_StepPlus_V6;   // Step structure
      SINI : Array[0..3] of USInt;
      LSTT : Array[0..7] of USInt;
      ATAJ : Array[0..7] of USInt;
      ATAB : Array[0..7] of USInt;
      PSTT : Array[0..7] of USInt;
      NSTT : Array[0..7] of USInt;
      ASSJ : Array[0..7] of USInt;
      ASSB : Array[0..7] of USInt;
      PTTS : Array[0..7] of USInt;
      NTTS : Array[0..7] of USInt;
      SW_SQTS : Array[0..7] of USInt;
      SWITCH : Array[0..1] of USInt;
      TVX : Array[0..3] of USInt;
      TTX : Array[0..3] of USInt;
      TSX : Array[0..3] of USInt;
      S00X : Array[0..3] of USInt;
      SOFFX : Array[0..3] of USInt;
      SONX : Array[0..3] of USInt;
      SAX : Array[0..3] of USInt;
      SERRX : Array[0..8] of USInt;
      SMX : Array[0..8] of USInt;
      S0X : Array[0..8] of USInt;
      S1X : Array[0..8] of USInt;
      IL_ALARM_INST : Diag_Alarm;
      SUP_ALARM_INST : Diag_Alarm;
      STEP_TIME_ALARM_INST : Diag_Alarm;
      IEC_TIMER_INST : IEC_TIMER;
      TRANSACTION_FLAG : Bool := false;
   END_VAR
   // SINI[0] := 2;
   // SINI[2] := 255;
   // SINI[3] := 255;
   // LSTT[0] := 255;
   // LSTT[1] := 255;
   // LSTT[2] := 255;
   // LSTT[3] := 255;
   // LSTT[4] := 255;
   // LSTT[5] := 1;
   // ATAJ[1] := 1;
   // ATAJ[2] := 2;
   // ATAJ[3] := 3;
   // ATAJ[4] := 4;
   // ATAJ[5] := 5;
   // ATAB[1] := 1;
   // ATAB[2] := 2;
   // ATAB[3] := 3;
   // ATAB[4] := 4;
   // ATAB[5] := 5;
   // PSTT[1] := 1;
   // PSTT[2] := 2;
   // PSTT[3] := 3;
   // PSTT[4] := 4;
   // PSTT[5] := 5;
   // NSTT[0] := 1;
   // NSTT[1] := 2;
   // NSTT[2] := 3;
   // NSTT[3] := 4;
   // NSTT[4] := 6;
   // NSTT[5] := 1;
   // ASSJ[1] := 1;
   // ASSJ[2] := 2;
   // ASSJ[3] := 3;
   // ASSJ[4] := 4;
   // ASSJ[5] := 5;
   // ASSB[1] := 1;
   // ASSB[2] := 5;
   // ASSB[3] := 3;
   // ASSB[4] := 4;
   // ASSB[5] := 2;
   // PTTS[0] := 255;
   // PTTS[2] := 1;
   // PTTS[3] := 2;
   // PTTS[4] := 3;
   // PTTS[5] := 1;
   // NTTS[1] := 1;
   // NTTS[2] := 2;
   // NTTS[3] := 3;
   // NTTS[4] := 4;
   // NTTS[5] := 5;
   // SW_SQTS[2] := 1;
   // SW_SQTS[3] := 1;
   // SW_SQTS[4] := 1;
   // SW_SQTS[5] := 2;
   // SWITCH[0] := 160;
   // TVX[0] := 16#1;
   // TTX[0] := 16#1;
   // TSX[0] := 16#1;
   // S00X[0] := 16#1;
   // SOFFX[0] := 16#1;
   // SONX[0] := 16#1;
   // SAX[0] := 16#1;
   // SERRX[0] := 16#1;
   // SMX[0] := 16#1;
   // S0X[0] := 16#1;
   // S1X[0] := 16#1;
   // LSTT[6] := 255;
   // ATAJ[6] := 6;
   // ATAB[6] := 6;
   // PSTT[6] := 6;
   // NSTT[6] := 7;
   // ASSJ[6] := 6;
   // ASSB[6] := 6;
   // PTTS[6] := 4;
   // NTTS[6] := 6;
   // SW_SQTS[6] := 1;
   // LSTT[7] := 1;
   // ATAJ[7] := 7;
   // ATAB[7] := 7;
   // PSTT[7] := 7;
   // NSTT[7] := 1;
   // ASSJ[7] := 7;
   // ASSB[7] := 7;
   // PTTS[7] := 6;
   // NTTS[7] := 7;
   // SW_SQTS[7] := 1;
BEGIN